HMI tags "Digitais"
   "Digitais_MB-01-YR" : Bool = PLC Digitais.MB-01-YR AT %DB300.DBX0.1, 1 s
   "Digitais_MB-01-YF" : Bool = PLC Digitais.MB-01-YF AT %DB300.DBX0.2, 1 s
   "Digitais_MB-01-YFF" : Bool = PLC Digitais.MB-01-YFF AT %DB300.DBX0.3, 1 s
   "Digitais_MB-01-MM" : Bool = PLC Digitais.MB-01-MM AT %DB300.DBX0.4, 1 s
   "Digitais_MB-01-MA" : Bool = PLC Digitais.MB-01-MA AT %DB300.DBX0.5, 1 s
   "Digitais_MB-01-EMER" : Bool = PLC Digitais.MB-01-EMER AT %DB300.DBX0.6, 1 s
   "Digitais_MB-01-MN" : Bool = PLC Digitais.MB-01-MN AT %DB300.DBX0.7, 1 s
   "Digitais_MB-01-ML" : Bool = PLC Digitais.MB-01-ML AT %DB300.DBX1.0, 1 s
   "Digitais_MB-01-YFI" : Bool = PLC Digitais.MB-01-YFI AT %DB300.DBX1.1, 1 s
   "Digitais_MB-01-YFA" : Bool = PLC Digitais.MB-01-YFA AT %DB300.DBX1.2, 1 s
   "Digitais_MB-01-YPTA" : Bool = PLC Digitais.MB-01-YPTA AT %DB300.DBX1.3, 1 s
   "Digitais_MB-01-HM" : Bool = PLC Digitais.MB-01-HM AT %DB300.DBX1.4, 1 s
   "Digitais_MB-01-RST" : Bool = PLC Digitais.MB-01-RST AT %DB300.DBX1.5, 1 s
   "Digitais_MB-01-INTRU" : Bool = PLC Digitais.MB-01-INTRU AT %DB300.DBX1.6, 1 s
   "Digitais_MB-01-YFB" : Bool = PLC Digitais.MB-01-YFB AT %DB300.DBX1.7, 1 s
   "Digitais_MB-02-YSH" : Bool = PLC Digitais.MB-02-YSH AT %DB300.DBX2.0, 1 s
   "Digitais_MB-02-YR" : Bool = PLC Digitais.MB-02-YR AT %DB300.DBX2.1, 1 s
   "Digitais_MB-02-YF" : Bool = PLC Digitais.MB-02-YF AT %DB300.DBX2.2, 1 s
   "Digitais_MB-02-YFF" : Bool = PLC Digitais.MB-02-YFF AT %DB300.DBX2.3, 1 s
   "Digitais_MB-02-MM" : Bool = PLC Digitais.MB-02-MM AT %DB300.DBX2.4, 1 s
   "Digitais_MB-02-MA" : Bool = PLC Digitais.MB-02-MA AT %DB300.DBX2.5, 1 s
   "Digitais_MB-02-EMER" : Bool = PLC Digitais.MB-02-EMER AT %DB300.DBX2.6, 1 s
   "Digitais_MB-02-MN" : Bool = PLC Digitais.MB-02-MN AT %DB300.DBX2.7, 1 s
   "Digitais_MB-02-ML" : Bool = PLC Digitais.MB-02-ML AT %DB300.DBX3.0, 1 s
   "Digitais_MB-02-YFI" : Bool = PLC Digitais.MB-02-YFI AT %DB300.DBX3.1, 1 s
   "Digitais_MB-02-YFA" : Bool = PLC Digitais.MB-02-YFA AT %DB300.DBX3.2, 1 s
   "Digitais_MB-02-YPTA" : Bool = PLC Digitais.MB-02-YPTA AT %DB300.DBX3.3, 1 s
   "Digitais_MB-02-HM" : Bool = PLC Digitais.MB-02-HM AT %DB300.DBX3.4, 1 s
   "Digitais_MB-02-RST" : Bool = PLC Digitais.MB-02-RST AT %DB300.DBX3.5, 1 s
   "Digitais_MB-02-INTRU" : Bool = PLC Digitais.MB-02-INTRU AT %DB300.DBX3.6, 1 s
   "Digitais_MB-02-YFB" : Bool = PLC Digitais.MB-02-YFB AT %DB300.DBX3.7, 1 s
   "Digitais_MB-03-YSH" : Bool = PLC Digitais.MB-03-YSH AT %DB300.DBX4.0, 1 s
   "Digitais_MB-03-YR" : Bool = PLC Digitais.MB-03-YR AT %DB300.DBX4.1, 1 s
   "Digitais_MB-03-YF" : Bool = PLC Digitais.MB-03-YF AT %DB300.DBX4.2, 1 s
   "Digitais_MB-03-YFF" : Bool = PLC Digitais.MB-03-YFF AT %DB300.DBX4.3, 1 s
   "Digitais_MB-03-MM" : Bool = PLC Digitais.MB-03-MM AT %DB300.DBX4.4, 1 s
   "Digitais_MB-03-MA" : Bool = PLC Digitais.MB-03-MA AT %DB300.DBX4.5, 1 s
   "Digitais_MB-03-EMER" : Bool = PLC Digitais.MB-03-EMER AT %DB300.DBX4.6, 1 s
   "Digitais_MB-03-MN" : Bool = PLC Digitais.MB-03-MN AT %DB300.DBX4.7, 1 s
   "Digitais_MB-03-ML" : Bool = PLC Digitais.MB-03-ML AT %DB300.DBX5.0, 1 s
   "Digitais_MB-03-YFI" : Bool = PLC Digitais.MB-03-YFI AT %DB300.DBX5.1, 1 s
   "Digitais_MB-03-YFA" : Bool = PLC Digitais.MB-03-YFA AT %DB300.DBX5.2, 1 s
   "Digitais_MB-03-YPTA" : Bool = PLC Digitais.MB-03-YPTA AT %DB300.DBX5.3, 1 s
   "Digitais_MB-03-HM" : Bool = PLC Digitais.MB-03-HM AT %DB300.DBX5.4, 1 s
   "Digitais_MB-03-RST" : Bool = PLC Digitais.MB-03-RST AT %DB300.DBX5.5, 1 s
   "Digitais_MB-03-INTRU" : Bool = PLC Digitais.MB-03-INTRU AT %DB300.DBX5.6, 1 s
   "Digitais_MB-03-YFB" : Bool = PLC Digitais.MB-03-YFB AT %DB300.DBX5.7, 1 s
   "Digitais_MB-04-YSH" : Bool = PLC Digitais.MB-04-YSH AT %DB300.DBX6.0, 1 s
   "Digitais_MB-04-YR" : Bool = PLC Digitais.MB-04-YR AT %DB300.DBX6.1, 1 s
   "Digitais_MB-04-YF" : Bool = PLC Digitais.MB-04-YF AT %DB300.DBX6.2, 1 s
   "Digitais_MB-04-YFF" : Bool = PLC Digitais.MB-04-YFF AT %DB300.DBX6.3, 1 s
   "Digitais_MB-04-MM" : Bool = PLC Digitais.MB-04-MM AT %DB300.DBX6.4, 1 s
   "Digitais_MB-04-MA" : Bool = PLC Digitais.MB-04-MA AT %DB300.DBX6.5, 1 s
   "Digitais_MB-04-EMER" : Bool = PLC Digitais.MB-04-EMER AT %DB300.DBX6.6, 1 s
   "Digitais_MB-04-MN" : Bool = PLC Digitais.MB-04-MN AT %DB300.DBX6.7, 1 s
   "Digitais_MB-04-ML" : Bool = PLC Digitais.MB-04-ML AT %DB300.DBX7.0, 1 s
   "Digitais_MB-04-YFI" : Bool = PLC Digitais.MB-04-YFI AT %DB300.DBX7.1, 1 s
   "Digitais_MB-04-YFA" : Bool = PLC Digitais.MB-04-YFA AT %DB300.DBX7.2, 1 s
   "Digitais_MB-04-YPTA" : Bool = PLC Digitais.MB-04-YPTA AT %DB300.DBX7.3, 1 s
   "Digitais_MB-04-HM" : Bool = PLC Digitais.MB-04-HM AT %DB300.DBX7.4, 1 s
   "Digitais_MB-04-RST" : Bool = PLC Digitais.MB-04-RST AT %DB300.DBX7.5, 1 s
   "Digitais_MB-04-INTRU" : Bool = PLC Digitais.MB-04-INTRU AT %DB300.DBX7.6, 1 s
   "Digitais_MB-04-YFB" : Bool = PLC Digitais.MB-04-YFB AT %DB300.DBX7.7, 1 s
   "Digitais_LIT_001-AL8" : Bool = PLC Digitais.LIT_001-AL8 AT %DB300.DBX8.0, 1 s
   "Digitais_LIT_001-AL9" : Bool = PLC Digitais.LIT_001-AL9 AT %DB300.DBX8.1, 1 s
   "Digitais_LIT_001-AL10" : Bool = PLC Digitais.LIT_001-AL10 AT %DB300.DBX8.2, 1 s
   "Digitais_LIT_001-AL11" : Bool = PLC Digitais.LIT_001-AL11 AT %DB300.DBX8.3, 1 s
   "Digitais_LIT_001-AL12" : Bool = PLC Digitais.LIT_001-AL12 AT %DB300.DBX8.4, 1 s
   "Digitais_LIT_001-AL13" : Bool = PLC Digitais.LIT_001-AL13 AT %DB300.DBX8.5, 1 s
   "Digitais_LIT_001-AL14" : Bool = PLC Digitais.LIT_001-AL14 AT %DB300.DBX8.6, 1 s
   "Digitais_LIT_001-AL15" : Bool = PLC Digitais.LIT_001-AL15 AT %DB300.DBX8.7, 1 s
   "Digitais_LIT_001-YHH" : Bool = PLC Digitais.LIT_001-YHH AT %DB300.DBX9.0, 1 s
   "Digitais_LIT_001-YH" : Bool = PLC Digitais.LIT_001-YH AT %DB300.DBX9.1, 1 s
   "Digitais_LIT_001-YL" : Bool = PLC Digitais.LIT_001-YL AT %DB300.DBX9.2, 1 s
   "Digitais_LIT_001-YLL" : Bool = PLC Digitais.LIT_001-YLL AT %DB300.DBX9.3, 1 s
   "Digitais_LIT_001-YFS" : Bool = PLC Digitais.LIT_001-YFS AT %DB300.DBX9.4, 1 s
   "Digitais_LIT_001-AL5" : Bool = PLC Digitais.LIT_001-AL5 AT %DB300.DBX9.5, 1 s
   "Digitais_LIT_001-AL6" : Bool = PLC Digitais.LIT_001-AL6 AT %DB300.DBX9.6, 1 s
   "Digitais_LIT_001-AL7" : Bool = PLC Digitais.LIT_001-AL7 AT %DB300.DBX9.7, 1 s
   "Digitais_PCM_EEE_EMER" : Bool = PLC Digitais.PCM_EEE_EMER AT %DB300.DBX10.0, 1 s
   "Digitais_PCM_EEE_K27" : Bool = PLC Digitais.PCM_EEE_K27 AT %DB300.DBX10.1, 1 s
   "Digitais_PCM_EEE_DISJ_LIG" : Bool = PLC Digitais.PCM_EEE_DISJ_LIG AT %DB300.DBX10.2, 1 s
   "Digitais_PCM_EEE_DISJ_DESLIG" : Bool = PLC Digitais.PCM_EEE_DISJ_DESLIG AT %DB300.DBX10.3, 1 s
   "Digitais_PCM_EEE_DISJ_YFAL" : Bool = PLC Digitais.PCM_EEE_DISJ_YFAL AT %DB300.DBX10.4, 1 s
   "Digitais_PCM_EEE_DISJ_FAL_GR" : Bool = PLC Digitais.PCM_EEE_DISJ_FAL_GR AT %DB300.DBX10.5, 1 s
   "Digitais_PCM_EEE_TR01_KA3" : Bool = PLC Digitais.PCM_EEE_TR01_KA3 AT %DB300.DBX10.6, 1 s
   "Digitais_PCM_EEE_TR01_KA4" : Bool = PLC Digitais.PCM_EEE_TR01_KA4 AT %DB300.DBX10.7, 1 s
   "Digitais_PCM_EEE_TR01_KA5" : Bool = PLC Digitais.PCM_EEE_TR01_KA5 AT %DB300.DBX11.0, 1 s
   "Digitais_PCM_EEE_INTRU" : Bool = PLC Digitais.PCM_EEE_INTRU AT %DB300.DBX11.1, 1 s
   "Digitais_PCM_EEE_RSERVA_0" : Bool = PLC Digitais.PCM_EEE_RSERVA_0 AT %DB300.DBX11.2, 1 s
   "Digitais_PCM_EEE_RSERVA_1" : Bool = PLC Digitais.PCM_EEE_RSERVA_1 AT %DB300.DBX11.3, 1 s
   "Digitais_PCM_EEE_RSERVA_2" : Bool = PLC Digitais.PCM_EEE_RSERVA_2 AT %DB300.DBX11.4, 1 s
   "Digitais_PCM_EEE_RSERVA_3" : Bool = PLC Digitais.PCM_EEE_RSERVA_3 AT %DB300.DBX11.5, 1 s
   "Digitais_PCM_EEE_RSERVA_4" : Bool = PLC Digitais.PCM_EEE_RSERVA_4 AT %DB300.DBX11.6, 1 s
   "Digitais_PCM_EEE_RSERVA_5" : Bool = PLC Digitais.PCM_EEE_RSERVA_5 AT %DB300.DBX11.7, 1 s
   "Digitais_QGBT_EMER" : Bool = PLC Digitais.QGBT_EMER AT %DB300.DBX12.0, 1 s
   "Digitais_QGBT_K27" : Bool = PLC Digitais.QGBT_K27 AT %DB300.DBX12.1, 1 s
   "Digitais_QGBT_DJL" : Bool = PLC Digitais.QGBT_DJL AT %DB300.DBX12.2, 1 s
   "Digitais_QGBT_DJD" : Bool = PLC Digitais.QGBT_DJD AT %DB300.DBX12.3, 1 s
   "Digitais_QGBT_DJYFAL" : Bool = PLC Digitais.QGBT_DJYFAL AT %DB300.DBX12.4, 1 s
   "Digitais_QGBT_INTRU" : Bool = PLC Digitais.QGBT_INTRU AT %DB300.DBX12.5, 1 s
   "Digitais_QGBT_RESERVA_0" : Bool = PLC Digitais.QGBT_RESERVA_0 AT %DB300.DBX12.6, 1 s
   "Digitais_QGBT_RESERVA_1" : Bool = PLC Digitais.QGBT_RESERVA_1 AT %DB300.DBX12.7, 1 s
   "Digitais_QGBT_RESERVA_2" : Bool = PLC Digitais.QGBT_RESERVA_2 AT %DB300.DBX13.0, 1 s
   "Digitais_QGBT_RESERVA_3" : Bool = PLC Digitais.QGBT_RESERVA_3 AT %DB300.DBX13.1, 1 s
   "Digitais_QGBT_RESERVA_4" : Bool = PLC Digitais.QGBT_RESERVA_4 AT %DB300.DBX13.2, 1 s
   "Digitais_QGBT_RESERVA_5" : Bool = PLC Digitais.QGBT_RESERVA_5 AT %DB300.DBX13.3, 1 s
   "Digitais_QGBT_RESERVA_6" : Bool = PLC Digitais.QGBT_RESERVA_6 AT %DB300.DBX13.4, 1 s
   "Digitais_QGBT_RESERVA_7" : Bool = PLC Digitais.QGBT_RESERVA_7 AT %DB300.DBX13.5, 1 s
   "Digitais_QGBT_RESERVA_8" : Bool = PLC Digitais.QGBT_RESERVA_8 AT %DB300.DBX13.6, 1 s
   "Digitais_QGBT_RESERVA_9" : Bool = PLC Digitais.QGBT_RESERVA_9 AT %DB300.DBX13.7, 1 s
   "Digitais_LSL_001" : Bool = PLC Digitais.LSL_001 AT %DB300.DBX14.0, 1 s
   "Digitais_LSH_001" : Bool = PLC Digitais.LSH_001 AT %DB300.DBX14.1, 1 s
   "Digitais_LSL_002" : Bool = PLC Digitais.LSL_002 AT %DB300.DBX14.2, 1 s
   "Digitais_LSH_002" : Bool = PLC Digitais.LSH_002 AT %DB300.DBX14.3, 1 s
   "Digitais_LS_RESERVA_0" : Bool = PLC Digitais.LS_RESERVA_0 AT %DB300.DBX14.4, 1 s
   "Digitais_LS_RESERVA_1" : Bool = PLC Digitais.LS_RESERVA_1 AT %DB300.DBX14.5, 1 s
   "Digitais_LS_RESERVA_2" : Bool = PLC Digitais.LS_RESERVA_2 AT %DB300.DBX14.6, 1 s
   "Digitais_LS_RESERVA_3" : Bool = PLC Digitais.LS_RESERVA_3 AT %DB300.DBX14.7, 1 s
   "Digitais_LS_RESERVA_4" : Bool = PLC Digitais.LS_RESERVA_4 AT %DB300.DBX15.0, 1 s
   "Digitais_LS_RESERVA_5" : Bool = PLC Digitais.LS_RESERVA_5 AT %DB300.DBX15.1, 1 s
   "Digitais_LS_RESERVA_6" : Bool = PLC Digitais.LS_RESERVA_6 AT %DB300.DBX15.2, 1 s
   "Digitais_LS_RESERVA_7" : Bool = PLC Digitais.LS_RESERVA_7 AT %DB300.DBX15.3, 1 s
   "Digitais_LS_RESERVA_8" : Bool = PLC Digitais.LS_RESERVA_8 AT %DB300.DBX15.4, 1 s
   "Digitais_LS_RESERVA_9" : Bool = PLC Digitais.LS_RESERVA_9 AT %DB300.DBX15.5, 1 s
   "Digitais_LS_RESERVA_10" : Bool = PLC Digitais.LS_RESERVA_10 AT %DB300.DBX15.6, 1 s
   "Digitais_LS_RESERVA_11" : Bool = PLC Digitais.LS_RESERVA_11 AT %DB300.DBX15.7, 1 s
   "Digitais_PCE_EEE_INTRU" : Bool = PLC Digitais.PCE_EEE_INTRU AT %DB300.DBX16.0, 1 s
   "Digitais_PCE_EEE_UPS_ALM" : Bool = PLC Digitais.PCE_EEE_UPS_ALM AT %DB300.DBX16.1, 1 s
   "Digitais_PCE_EEE_UPS_FE" : Bool = PLC Digitais.PCE_EEE_UPS_FE AT %DB300.DBX16.2, 1 s
   "Digitais_PCE_EEE_UPS_CHAR" : Bool = PLC Digitais.PCE_EEE_UPS_CHAR AT %DB300.DBX16.3, 1 s
   "Digitais_PCM-E-CF-01-P100-YFC" : Bool = PLC Digitais.PCM-E-CF-01-P100-YFC AT %DB300.DBX16.4, 1 s
   "Digitais_QGBT-AUX-01-P100-YFC" : Bool = PLC Digitais.QGBT-AUX-01-P100-YFC AT %DB300.DBX16.5, 1 s

HMI tags "Setpoints"
   "SETPOINTS_MB-01-SP" : Real = PLC SETPOINTS.MB-01-SP AT %DB305.DBD0, 1 s
   "SETPOINTS_MB-02-SP" : Real = PLC SETPOINTS.MB-02-SP AT %DB305.DBD4, 1 s
   "SETPOINTS_MB-03-SP" : Real = PLC SETPOINTS.MB-03-SP AT %DB305.DBD8, 1 s
   "SETPOINTS_MB-04-SP" : Real = PLC SETPOINTS.MB-04-SP AT %DB305.DBD12, 1 s
   "SETPOINTS_LIT_001-SPHH" : Real = PLC SETPOINTS.LIT_001-SPHH AT %DB305.DBD16, 1 s
   "SETPOINTS_LIT_001-SPH" : Real = PLC SETPOINTS.LIT_001-SPH AT %DB305.DBD20, 1 s
   "SETPOINTS_LIT_001-SPL" : Real = PLC SETPOINTS.LIT_001-SPL AT %DB305.DBD24, 1 s
   "SETPOINTS_LIT_001-SPLL" : Real = PLC SETPOINTS.LIT_001-SPLL AT %DB305.DBD28, 1 s
   "SETPOINTS_LIT_001-SPM" : Real = PLC SETPOINTS.LIT_001-SPM AT %DB305.DBD32, 1 s
   "SETPOINTS_LIT_001-SPC" : Real = PLC SETPOINTS.LIT_001-SPC AT %DB305.DBD36, 1 s
   "SETPOINTS_LIT-001-P" : Real = PLC SETPOINTS.LIT-001-P AT %DB305.DBD40, 1 s
   "SETPOINTS_SP_NVL_MIN" : Real = PLC SETPOINTS.SP_NVL_MIN AT %DB305.DBD44, 1 s
   "SETPOINTS_MB-P-SP-DL" : Real = PLC SETPOINTS.MB-P-SP-DL AT %DB305.DBD48, 1 s
   "SETPOINTS_MB-P-SP-L" : Real = PLC SETPOINTS.MB-P-SP-L AT %DB305.DBD52, 1 s
   "SETPOINTS_MB-C1-SP-DL" : Real = PLC SETPOINTS.MB-C1-SP-DL AT %DB305.DBD56, 1 s
   "SETPOINTS_MB-C1-SP-L" : Real = PLC SETPOINTS.MB-C1-SP-L AT %DB305.DBD60, 1 s
   "SETPOINTS_MB-C2-SP-DL" : Real = PLC SETPOINTS.MB-C2-SP-DL AT %DB305.DBD64, 1 s
   "SETPOINTS_MB-C2-SP-L" : Real = PLC SETPOINTS.MB-C2-SP-L AT %DB305.DBD68, 1 s
   "SETPOINTS_MB-C3-SP-DL" : Real = PLC SETPOINTS.MB-C3-SP-DL AT %DB305.DBD72, 1 s
   "SETPOINTS_MB-C3-SP-L" : Real = PLC SETPOINTS.MB-C3-SP-L AT %DB305.DBD76, 1 s

HMI tags "Variaveis"
   "VARIAVEIS_MB-01-YST" : Real = PLC VARIAVEIS.MB-01-YST AT %DB304.DBD0, 1 s
   "VARIAVEIS_MB-01-YIT" : Real = PLC VARIAVEIS.MB-01-YIT AT %DB304.DBD4, 1 s
   "VARIAVEIS_MB-02-YIT" : Real = PLC VARIAVEIS.MB-02-YIT AT %DB304.DBD8, 1 s
   "VARIAVEIS_MB-02-YST" : Real = PLC VARIAVEIS.MB-02-YST AT %DB304.DBD12, 1 s
   "VARIAVEIS_MB-03-YIT" : Real = PLC VARIAVEIS.MB-03-YIT AT %DB304.DBD16, 1 s
   "VARIAVEIS_MB-03-YST" : Real = PLC VARIAVEIS.MB-03-YST AT %DB304.DBD20, 1 s
   "VARIAVEIS_MB-04-YIT" : Real = PLC VARIAVEIS.MB-04-YIT AT %DB304.DBD24, 1 s
   "VARIAVEIS_MB-04-YST" : Real = PLC VARIAVEIS.MB-04-YST AT %DB304.DBD28, 1 s
   "VARIAVEIS_LIT_001" : Real = PLC VARIAVEIS.LIT_001 AT %DB304.DBD32, 1 s
   "VARIAVEIS_LIT_001-P" : Real = PLC VARIAVEIS.LIT_001-P AT %DB304.DBD36, 1 s
   "VARIAVEIS_PCM-E-CF-01-04-P100-ETRS" : Real = PLC VARIAVEIS.PCM-E-CF-01-04-P100-ETRS AT %DB304.DBD40, 1 s
   "VARIAVEIS_PCM-E-CF-01-04-P100-ETST" : Real = PLC VARIAVEIS.PCM-E-CF-01-04-P100-ETST AT %DB304.DBD44, 1 s
   "VARIAVEIS_PCM-E-CF-01-04-P100-ETTR" : Real = PLC VARIAVEIS.PCM-E-CF-01-04-P100-ETTR AT %DB304.DBD48, 1 s
   "VARIAVEIS_PCM-E-CF-01-04-P100-ITR" : Real = PLC VARIAVEIS.PCM-E-CF-01-04-P100-ITR AT %DB304.DBD52, 1 s
   "VARIAVEIS_PCM-E-CF-01-04-P100-ITS" : Real = PLC VARIAVEIS.PCM-E-CF-01-04-P100-ITS AT %DB304.DBD56, 1 s
   "VARIAVEIS_PCM-E-CF-01-04-P100-ITT" : Real = PLC VARIAVEIS.PCM-E-CF-01-04-P100-ITT AT %DB304.DBD60, 1 s
   "VARIAVEIS_PCM-E-CF-01-04-P100-JPT" : Real = PLC VARIAVEIS.PCM-E-CF-01-04-P100-JPT AT %DB304.DBD64, 1 s
   "VARIAVEIS_PCM-E-CF-01-04-P100-JQT" : Real = PLC VARIAVEIS.PCM-E-CF-01-04-P100-JQT AT %DB304.DBD68, 1 s
   "VARIAVEIS_PCM-E-CF-01-04-P100-JST" : Real = PLC VARIAVEIS.PCM-E-CF-01-04-P100-JST AT %DB304.DBD72, 1 s
   "VARIAVEIS_PCM-E-CF-01-04-P100-FP" : Real = PLC VARIAVEIS.PCM-E-CF-01-04-P100-FP AT %DB304.DBD76, 1 s
   "VARIAVEIS_QGBT-AUX-01-P100-ETRS" : Real = PLC VARIAVEIS.QGBT-AUX-01-P100-ETRS AT %DB304.DBD80, 1 s
   "VARIAVEIS_QGBT-AUX-01-P100-ETST" : Real = PLC VARIAVEIS.QGBT-AUX-01-P100-ETST AT %DB304.DBD84, 1 s
   "VARIAVEIS_QGBT-AUX-01-P100-ETTR" : Real = PLC VARIAVEIS.QGBT-AUX-01-P100-ETTR AT %DB304.DBD88, 1 s
   "VARIAVEIS_QGBT-AUX-01-P100-ITR" : Real = PLC VARIAVEIS.QGBT-AUX-01-P100-ITR AT %DB304.DBD92, 1 s
   "VARIAVEIS_QGBT-AUX-01-P100-ITS" : Real = PLC VARIAVEIS.QGBT-AUX-01-P100-ITS AT %DB304.DBD96, 1 s
   "VARIAVEIS_QGBT-AUX-01-P100-ITT" : Real = PLC VARIAVEIS.QGBT-AUX-01-P100-ITT AT %DB304.DBD100, 1 s
   "VARIAVEIS_QGBT-AUX-01-P100-JPT" : Real = PLC VARIAVEIS.QGBT-AUX-01-P100-JPT AT %DB304.DBD104, 1 s
   "VARIAVEIS_QGBT-AUX-01-P100-JQT" : Real = PLC VARIAVEIS.QGBT-AUX-01-P100-JQT AT %DB304.DBD108, 1 s
   "VARIAVEIS_QGBT-AUX-01-P100-JST" : Real = PLC VARIAVEIS.QGBT-AUX-01-P100-JST AT %DB304.DBD112, 1 s
   "VARIAVEIS_QGBT-AUX-01-P100-FP" : Real = PLC VARIAVEIS.QGBT-AUX-01-P100-FP AT %DB304.DBD116, 1 s

HMI tags "STATUS"
   "STATUS_MB-01-YSP" : Bool = PLC STATUS.MB-01-YSP AT %DB302.DBX0.6, 1 s
   "STATUS_MB-02-YSP" : Bool = PLC STATUS.MB-02-YSP AT %DB302.DBX0.7, 1 s
   "STATUS_MB-03-YSP" : Bool = PLC STATUS.MB-03-YSP AT %DB302.DBX1.1, 1 s
   "STATUS_MB-01-YC1" : Bool = PLC STATUS.MB-01-YC1 AT %DB302.DBX1.2, 1 s
   "STATUS_MB-02-YC1" : Bool = PLC STATUS.MB-02-YC1 AT %DB302.DBX1.3, 1 s
   "STATUS_MB-03-YC1" : Bool = PLC STATUS.MB-03-YC1 AT %DB302.DBX1.5, 1 s
   "STATUS_MB-01-YC2" : Bool = PLC STATUS.MB-01-YC2 AT %DB302.DBX1.6, 1 s
   "STATUS_MB-02-YC2" : Bool = PLC STATUS.MB-02-YC2 AT %DB302.DBX1.7, 1 s
   "STATUS_MB-03-YC2" : Bool = PLC STATUS.MB-03-YC2 AT %DB302.DBX2.1, 1 s
   "STATUS_MB-04-YSP" : Bool = PLC STATUS.MB-04-YSP AT %DB302.DBX1.0, 1 s
   "STATUS_MB-04-YC1" : Bool = PLC STATUS.MB-04-YC1 AT %DB302.DBX1.4, 1 s
   "STATUS_MB-04-YC2" : Bool = PLC STATUS.MB-04-YC2 AT %DB302.DBX2.0, 1 s

discrete alarms
   1: 'Elevatoria principal 1 falha', class Errors, trigger "ALM0" bit 10
   2: 'Elevatoria principal 1 falta de fase', class Errors, trigger "ALM0" bit 11
   3: 'Elevatoria principal 1 emergencia', class Errors, trigger "ALM0" bit 14
   5: 'Elevatoria principal 1 com falha no inversor', class Errors, trigger "ALM0" bit 1
   6: 'Elevatoria principal 1 com falha no acionamento', class Errors, trigger "ALM0" bit 2
   7: 'Elevatoria principal 1 com proteção térmica atuada', class Errors, trigger "ALM0" bit 3
   8: 'Elevatoria principal 1 intrusão no painel', class Errors, trigger "ALM0" bit 6
   9: 'Elevatoria principal 1 defeito na bomba', class Errors, trigger "ALM0" bit 7
   10: 'Elevatoria principal 2 falha', class Errors, trigger "ALM2" bit 10
   11: 'Elevatoria principal 2 falta de fase', class Errors, trigger "ALM2" bit 11
   12: 'Elevatoria principal 2 emergencia', class Errors, trigger "ALM2" bit 14
   14: 'Elevatoria principal 2 com falha no inversor', class Errors, trigger "ALM2" bit 1
   15: 'Elevatoria principal 2 com falha no acionamento', class Errors, trigger "ALM2" bit 2
   16: 'Elevatoria principal 2 com proteção térmica atuada', class Errors, trigger "ALM2" bit 3
   17: 'Elevatoria principal 2 intrusão no painel', class Errors, trigger "ALM2" bit 6
   18: 'Elevatoria principal 2 defeito na bomba', class Errors, trigger "ALM2" bit 7
   19: 'Elevatoria principal 3 falha', class Errors, trigger "ALM4" bit 10
   20: 'Elevatoria principal 3 falta de fase', class Errors, trigger "ALM4" bit 11
   21: 'Elevatoria principal 3 emergencia', class Errors, trigger "ALM4" bit 14
   23: 'Elevatoria principal 3 com falha no inversor', class Errors, trigger "ALM4" bit 1
   24: 'Elevatoria principal 3 com falha no acionamento', class Errors, trigger "ALM4" bit 2
   25: 'Elevatoria principal 3 com proteção térmica atuada', class Errors, trigger "ALM4" bit 3
   26: 'Elevatoria principal 3 intrusão no painel', class Errors, trigger "ALM4" bit 6
   27: 'Elevatoria principal 3 defeito na bomba', class Errors, trigger "ALM4" bit 7
   28: 'Elevatoria principal 4 falha', class Errors, trigger "ALM6" bit 10
   29: 'Elevatoria principal 4 falta de fase', class Errors, trigger "ALM6" bit 11
   30: 'Elevatoria principal 4 emergencia', class Errors, trigger "ALM6" bit 14
   32: 'Elevatoria principal 4 com falha no inversor', class Errors, trigger "ALM6" bit 1
   33: 'Elevatoria principal 4 com falha no acionamento', class Errors, trigger "ALM6" bit 2
   34: 'Elevatoria principal 4 com proteção térmica atuada', class Errors, trigger "ALM6" bit 3
   35: 'Elevatoria principal 4 intrusão no painel', class Errors, trigger "ALM6" bit 6
   36: 'Elevatoria principal 4 defeito na bomba', class Errors, trigger "ALM6" bit 7
   37: 'Alarme de nível muito alto do tanque', class Errors, trigger "ALM8" bit 0
   38: 'Alarme de nível alto do tanque', class Errors, trigger "ALM8" bit 1
   39: 'Alarme de nível baixo do tanque', class Errors, trigger "ALM8" bit 2
   40: 'Alarme de nível muito baixo do tanque', class Errors, trigger "ALM8" bit 3
   41: 'Transmissor de nível do tanque com falha de sinal', class Errors, trigger "ALM8" bit 4
   42: 'PCM-E-CF-01-04 BOTAO DE EMERGENCIA - ATUADO', class Errors, trigger "ALM10" bit 8
   43: 'PCM-E-CF-01-04 RELE DE PROTECAO FUNCAO 27 - ATUADO', class Errors, trigger "ALM10" bit 9
   44: 'PCM-E-CF-01-04 DISJUNTOR GERAL STATUS - FALHA', class Errors, trigger "ALM10" bit 12
   45: 'PCM-E-CF-01-04 FALHA GERAL ATUADO', class Errors, trigger "ALM10" bit 13
   46: 'PCM-E-CF-01-04 TRANSFORMADOR -TR-01 ALARME TEMP 150°', class Errors, trigger "ALM10" bit 14
   47: 'PCM-E-CF-01-04 TRANSFORMADOR -TR-01 ALARME TEMP 155°', class Errors, trigger "ALM10" bit 15
   48: 'PCM-E-CF-01-04 TRANSFORMADOR -TR-01 FALHA PROTECAO', class Errors, trigger "ALM10" bit 0
   49: 'PCM-E-CF-01-04 INTRUSAO NO PAINEL (COLUNA 01~04)', class Errors, trigger "ALM10" bit 1
   50: 'QGBT-AUX-01 BOTAO DE EMERGENCIA ATUADO', class Errors, trigger "ALM12" bit 8
   51: 'QGBT-AUX-01 RELE DE PROTECAO FUNCAO 27/59 ATUADO', class Errors, trigger "ALM12" bit 9
   52: 'QGBT-AUX-01 DISJUNTOR GERAL FALHA - TRIP', class Errors, trigger "ALM12" bit 12
   53: 'QGBT-AUX-01 INTRUSAO NO PAINEL', class Errors, trigger "ALM12" bit 13
   54: 'INTRUSAO NO PAINEL', class Errors, trigger "ALM16" bit 8
   55: 'UPS EM ALARME FALHA NA BATERIA', class Errors, trigger "ALM16" bit 9
   56: 'UPS EM OPERACAO FALTA DE ENERGIA', class Errors, trigger "ALM16" bit 10
   57: 'UPS EM ALARME BATERIA CARREGADA', class Errors, trigger "ALM16" bit 11

screen "EEEB" 800x480, template "Template_1"
   GraphicView "Template_Graphic view_3" at 143,92 size 589x312; Picture "EEEB_2"
   Bar "Bar_1" at 679,137 size 57x267; MinimumValue 0; MaximumValue 100
      ProcessValue <- "VARIAVEIS_LIT_001-P"
   GraphicView "Graphic view_1" at 280,337 size 47x47; Picture "Submersa_vm"
      Visibility <- "Digitais_MB-01-YSH"
   GraphicView "Graphic view_2" at 280,337 size 47x47; Picture "Submersa_am"
      Visibility <- "Digitais_MB-01-YF"
   GraphicView "Graphic view_3" at 280,337 size 47x47; Picture "Submersa_azul"
      Visibility <- "COMANDOS_MB-01-HS7"
   GraphicView "Graphic view_4" at 395,337 size 47x47; Picture "Submersa_vm"
      Visibility <- "Digitais_MB-02-YSH"
   GraphicView "Graphic view_5" at 395,337 size 47x47; Picture "Submersa_am"
      Visibility <- "Digitais_MB-02-YF"
   GraphicView "Graphic view_6" at 395,337 size 47x47; Picture "Submersa_azul"
      Visibility <- "COMANDOS_MB-02-HS7"
   GraphicView "Graphic view_7" at 510,337 size 47x47; Picture "Submersa_vm"
      Visibility <- "Digitais_MB-03-YSH"
   GraphicView "Graphic view_8" at 510,337 size 47x47; Picture "Submersa_am"
      Visibility <- "Digitais_MB-03-YF"
   GraphicView "Graphic view_9" at 510,337 size 47x47; Picture "Submersa_azul"
      Visibility <- "COMANDOS_MB-03-HS7"
   TextField "Text field_1" at 286,384 size 29x14; Text 'MB-01'
   TextField "Text field_2" at 403,384 size 29x14; Text 'MB-02'
   TextField "Text field_3" at 517,384 size 29x14; Text 'MB-03'
   TextField "Text field_4" at 248,328 size 25x16; Text 'AUT'
      Visibility <- "COMANDOS_MB-01-HS1"
   TextField "Text field_5" at 248,345 size 25x16; Text 'REM'
      Visibility <- "Digitais_MB-01-YR"
   TextField "Text field_6" at 296,322 size 25x16; Text 'P'
      Visibility <- "STATUS_MB-01-YSP"
   TextField "Text field_7" at 296,322 size 25x16; Text 'C1'
      Visibility <- "STATUS_MB-01-YC1"
   TextField "Text field_8" at 296,322 size 25x16; Text 'C2'
      Visibility <- "STATUS_MB-01-YC2"
   IOField "I/O field_3" at 222,363 size 54x17; FormatPattern 99.9; Unit  HZ
      ProcessValue <- "VARIAVEIS_MB-01-YST"
   IOField "I/O field_4" at 223,380 size 55x17; FormatPattern 999.9; Unit  A
      ProcessValue <- "VARIAVEIS_MB-01-YIT"
   TextField "Text field_9" at 364,328 size 25x16; Text 'AUT'
      Visibility <- "COMANDOS_MB-02-HS1"
   TextField "Text field_10" at 364,345 size 25x16; Text 'REM'
      Visibility <- "Digitais_MB-02-YR"
   TextField "Text field_11" at 412,322 size 25x16; Text 'P'
      Visibility <- "STATUS_MB-02-YSP"
   TextField "Text field_12" at 412,322 size 25x16; Text 'C1'
      Visibility <- "STATUS_MB-02-YC1"
   TextField "Text field_13" at 412,322 size 25x16; Text 'C2'
      Visibility <- "STATUS_MB-02-YC2"
   IOField "I/O field_5" at 338,363 size 54x17; FormatPattern 99.9; Unit  HZ
      ProcessValue <- "VARIAVEIS_MB-02-YST"
   IOField "I/O field_6" at 339,380 size 55x17; FormatPattern 999.9; Unit  A
      ProcessValue <- "VARIAVEIS_MB-02-YIT"
   TextField "Text field_14" at 478,328 size 25x16; Text 'AUT'
      Visibility <- "COMANDOS_MB-03-HS1"
   TextField "Text field_15" at 478,345 size 25x16; Text 'REM'
      Visibility <- "Digitais_MB-03-YR"
   TextField "Text field_16" at 526,322 size 25x16; Text 'P'
      Visibility <- "STATUS_MB-03-YSP"
   TextField "Text field_17" at 526,322 size 25x16; Text 'C1'
      Visibility <- "STATUS_MB-03-YC1"
   TextField "Text field_18" at 526,322 size 25x16; Text 'C2'
      Visibility <- "STATUS_MB-03-YC2"
   IOField "I/O field_7" at 452,363 size 54x17; FormatPattern 99.9; Unit  HZ
      ProcessValue <- "VARIAVEIS_MB-03-YST"
   IOField "I/O field_8" at 453,380 size 55x17; FormatPattern 999.9; Unit  A
      ProcessValue <- "VARIAVEIS_MB-03-YIT"
   IOField "I/O field_14" at 738,164 size 59x17; FormatPattern 99.99; Unit  m
      ProcessValue <- "VARIAVEIS_LIT_001"
      Appearance <- "Digitais_LIT_001-YFS"
   IOField "I/O field_17" at 738,180 size 59x17; FormatPattern 999.9; Unit  %
      ProcessValue <- "VARIAVEIS_LIT_001-P"
      Appearance <- "Digitais_LIT_001-YFS"
   TextField "Text field_19" at 772,148 size 25x16; Text 'HH'
      Visibility <- "Digitais_LIT_001-YHH"
   TextField "Text field_20" at 738,148 size 25x16; Text 'LL'
      Visibility <- "Digitais_LIT_001-YLL"
   TextField "Text field_21" at 738,197 size 25x16; Text 'L'
      Visibility <- "Digitais_LIT_001-YL"
   TextField "Text field_22" at 772,197 size 25x16; Text 'H'
      Visibility <- "Digitais_LIT_001-YH"
   Button "Button_5" at 332,10 size 96x32; TextOff 'pause loop'
      on Click: InvertBit("pause")
      Appearance <- "pause"
   IOField "I/O field_18" at 352,48 size 59x17; FormatPattern s99999
      ProcessValue <- "DIVERSOS_Looping"
      Visibility <- "pause"
   IOField "I/O field_1" at 567,363 size 54x17; FormatPattern 99.9; Unit  HZ
      ProcessValue <- "VARIAVEIS_MB-04-YST"
   IOField "I/O field_2" at 568,380 size 55x17; FormatPattern 999.9; Unit  A
      ProcessValue <- "VARIAVEIS_MB-04-YIT"
   TextField "Text field_23" at 646,322 size 25x16; Text 'P'
      Visibility <- "STATUS_MB-04-YSP"
   TextField "Text field_24" at 646,322 size 25x16; Text 'C1'
      Visibility <- "STATUS_MB-04-YC1"
   TextField "Text field_25" at 646,322 size 25x16; Text 'C2'
      Visibility <- "STATUS_MB-04-YC2"
   TextField "Text field_26" at 596,328 size 25x16; Text 'AUT'
      Visibility <- "COMANDOS_MB-04-HS1"
   TextField "Text field_27" at 596,345 size 25x16; Text 'REM'
      Visibility <- "Digitais_MB-04-YR"
   TextField "Text field_28" at 631,384 size 29x14; Text 'MB-04'
   GraphicView "Graphic view_10" at 624,337 size 47x47; Picture "Submersa_vm"
      Visibility <- "Digitais_MB-04-YSH"
   GraphicView "Graphic view_11" at 624,337 size 47x47; Picture "Submersa_am"
      Visibility <- "Digitais_MB-04-YF"
   GraphicView "Graphic view_12" at 624,337 size 47x47; Picture "Submersa_azul"
      Visibility <- "COMANDOS_MB-04-HS7"
   TextField "Text field_29" at 175,148 size 25x16; Text 'HH'
      Visibility <- "Digitais_LSH_002"
   TextField "Text field_30" at 175,378 size 25x16; Text 'LL'
      Visibility <- "Digitais_LSL_002"
   TextField "Text field_31" at 175,337 size 25x16; Text 'L'
      Visibility <- "Digitais_LSL_001"
   TextField "Text field_32" at 175,189 size 25x16; Text 'H'
      Visibility <- "Digitais_LSH_001"
   TextField "Text field_33" at 216,310 size 65x18; Text 'Manuteção'
      Visibility <- "Digitais_MB-01-MM"
   TextField "Text field_34" at 249,310 size 32x18; Text 'Local'
      Visibility <- "Digitais_MB-01-ML"
   TextField "Text field_35" at 217,310 size 64x18; Text 'Emegência'
      Visibility <- "Digitais_MB-01-EMER"
   TextField "Text field_36" at 331,310 size 65x18; Text 'Manuteção'
      Visibility <- "Digitais_MB-02-MM"
   TextField "Text field_37" at 364,310 size 32x18; Text 'Local'
      Visibility <- "Digitais_MB-02-ML"
   TextField "Text field_38" at 332,310 size 64x18; Text 'Emegência'
      Visibility <- "Digitais_MB-02-EMER"
   TextField "Text field_39" at 446,310 size 65x18; Text 'Manuteção'
      Visibility <- "Digitais_MB-03-MM"
   TextField "Text field_40" at 479,310 size 32x18; Text 'Local'
      Visibility <- "Digitais_MB-03-ML"
   TextField "Text field_41" at 447,310 size 64x18; Text 'Emegência'
      Visibility <- "Digitais_MB-03-EMER"
   TextField "Text field_42" at 561,310 size 65x18; Text 'Manuteção'
      Visibility <- "Digitais_MB-04-MM"
   TextField "Text field_43" at 594,310 size 32x18; Text 'Local'
      Visibility <- "Digitais_MB-04-ML"
   TextField "Text field_44" at 562,310 size 64x18; Text 'Emegência'
      Visibility <- "Digitais_MB-04-EMER"
   TextField "Text field_45" at 391,406 size 138x22; Text 'Emegência Acionado'
      Visibility <- "Digitais_PCM_EEE_EMER"

Template "Template_1" 800x480
   Button "Exit" at 724,444 size 50x36; TextOn 'Exit'; TextOff 'Exit'; PictureOn "ExitRuntime_KTP400_Basic_PN_TR"; PictureOff "SB_ExitRuntime_80x60_256c"
      on Release: StopRuntime(0)
   Button "Alarms" at 524,444 size 50x36; TextOn 'Alarms'; TextOff 'Alarms'; PictureOn "AlarmDisplay_KTP400_Basic_PN_TR"; PictureOff "AlarmDisplay_KTP400_Basic_PN_TR"
      on Release: function_ef3f5d25("Alarm window_1", -1)
   SymbolicIOField "Symbolic_IO_Field_Screen" at 185,7 size 510x49; TextOn '1'; TextOff '0'; TextList "TextList_ScreenNames"
      on Change: ActivateScreenByNumber("Tag_ScreenNumber", 0)
      ProcessValue <- "Tag_ScreenNumber"
   DateTimeField "HmiScreenItemData" at 695,29 size 102x22
   DateTimeField "HmiScreenItemData_1" at 686,5 size 111x22
   Group "Group" at 0,0 size 179x67; Picture "consbem"
   Button "Start screen_1" at 26,444 size 50x36; TextOn 'EEEB / Start screen'; TextOff 'EEEB / Start screen'; PictureOn "NavigateHome_KTP400_Basic_PN_TR"; PictureOff "NavigateHome_KTP400_Basic_PN_TR"
      on Release: ActivateScreen("EEEB", 1)
   Button "Start screen_2" at 125,444 size 50x36; TextOn 'Ajustes / Start screen'; TextOff 'Ajustes / Start screen'; PictureOn "NavigateHome_KTP400_Basic_PN_TR"; PictureOff "NavigateHome_KTP400_Basic_PN_TR"
      on Release: ActivateScreen("Ajustes", 1)
   Button "Start screen_3" at 226,444 size 50x36; TextOn 'Comando / Start screen'; TextOff 'Comando / Start screen'; PictureOn "NavigateHome_KTP400_Basic_PN_TR"; PictureOff "NavigateHome_KTP400_Basic_PN_TR"
      on Release: ActivateScreen("Comandos", 1)
   Button "Start screen_4" at 328,444 size 50x36; TextOn 'PID / Start screen'; TextOff 'PID / Start screen'; PictureOn "NavigateHome_KTP400_Basic_PN_TR"; PictureOff "NavigateHome_KTP400_Basic_PN_TR"
      on Release: ActivateScreen("PID", 1)
   Button "Start screen_5" at 426,444 size 50x36; TextOn 'Monitor. / Start screen'; TextOff 'Monitor. / Start screen'; PictureOn "NavigateHome_KTP400_Basic_PN_TR"; PictureOff "NavigateHome_KTP400_Basic_PN_TR"
      on Release: ActivateScreen("Monitoramento", 1)
   Softkey "Softkey_F1" at 0,0 size 0x0
      on KeyUp: ActivateScreen("EEEB", 0)
   Softkey "Softkey_F2" at 0,0 size 0x0
      on KeyUp: ActivateScreen("Ajustes", 1)
   Softkey "Softkey_F3" at 0,0 size 0x0
      on KeyUp: ActivateScreen("Comandos", 0)
   Softkey "Softkey_F4" at 0,0 size 0x0
      on KeyUp: ActivateScreen("PID", 1)
   GraphicView "Template_Graphic view_2" at 60,0 size 60x67; Picture "Consbem_novo"
   GraphicView "Template_Graphic view_3" at 119,0 size 60x67; Picture "logo-saae-header"
   GraphicView "Template_Graphic view_4" at 0,0 size 60x67; Picture "logo cápua"
   Softkey "Softkey_F5" at 0,0 size 0x0
      on KeyUp: ActivateScreen("Monitoramento", 0)
   Softkey "Softkey_F6" at 0,0 size 0x0
      on KeyUp: function_ef3f5d25("Alarm window_1", -1)

screen "Monitoramento" 800x480, template "Template_1"
   IOField "I/O field_9" at 649,330 size 71x17; FormatPattern 999.99; Unit  kW
      ProcessValue <- "VARIAVEIS_QGBT-AUX-01-P100-JPT"
      Appearance <- "Digitais_LIT_001-YFS"
   TextField "Text field_14" at 607,295 size 78x23; Text 'Potências'
   TextField "Text field_15" at 604,327 size 40x20; Text 'Ativa'
   IOField "I/O field_10" at 649,352 size 71x17; FormatPattern 999.99; Unit  KVA
      ProcessValue <- "VARIAVEIS_QGBT-AUX-01-P100-JST"
      Appearance <- "Digitais_LIT_001-YFS"
   TextField "Text field_16" at 577,349 size 67x20; Text 'Aparente'
   IOField "I/O field_11" at 649,374 size 71x17; FormatPattern 999.99
      ProcessValue <- "VARIAVEIS_QGBT-AUX-01-P100-FP"
      Appearance <- "Digitais_LIT_001-YFS"
   TextField "Text field_17" at 525,371 size 119x20; Text 'Fator de Potência'
   IOField "I/O field_12" at 423,330 size 71x17; FormatPattern 999.99; Unit  A
      ProcessValue <- "VARIAVEIS_QGBT-AUX-01-P100-ITR"
      Appearance <- "Digitais_LIT_001-YFS"
   TextField "Text field_18" at 380,295 size 79x23; Text 'Correntes'
   TextField "Text field_19" at 370,327 size 47x20; Text 'Fase R'
   IOField "I/O field_13" at 423,352 size 71x17; FormatPattern 999.99; Unit  A
      ProcessValue <- "VARIAVEIS_QGBT-AUX-01-P100-ITS"
      Appearance <- "Digitais_LIT_001-YFS"
   TextField "Text field_20" at 371,349 size 46x20; Text 'Fase S'
   IOField "I/O field_15" at 423,374 size 71x17; FormatPattern 999.99; Unit  A
      ProcessValue <- "VARIAVEIS_QGBT-AUX-01-P100-ITT"
      Appearance <- "Digitais_LIT_001-YFS"
   TextField "Text field_21" at 372,371 size 45x20; Text 'Fase T'
   IOField "I/O field_16" at 202,330 size 71x17; FormatPattern 999.99; Unit  V
      ProcessValue <- "VARIAVEIS_QGBT-AUX-01-P100-ETRS"
      Appearance <- "Digitais_LIT_001-YFS"
   TextField "Text field_22" at 166,295 size 66x23; Text 'Tensões'
   TextField "Text field_23" at 133,327 size 63x20; Text 'Fase R/S'
   IOField "I/O field_17" at 202,352 size 71x17; FormatPattern 999.99; Unit  V
      ProcessValue <- "VARIAVEIS_QGBT-AUX-01-P100-ETST"
      Appearance <- "Digitais_LIT_001-YFS"
   TextField "Text field_24" at 133,349 size 61x20; Text 'Fase S/T'
   IOField "I/O field_18" at 202,374 size 71x17; FormatPattern 999.99; Unit  V
      ProcessValue <- "VARIAVEIS_QGBT-AUX-01-P100-ETTR"
      Appearance <- "Digitais_LIT_001-YFS"
   TextField "Text field_25" at 133,371 size 62x20; Text 'Fase T/R'
   TextField "Text field_26" at 350,263 size 120x23; Text 'QGBT-AUX-01'
   IOField "I/O field_6" at 649,154 size 71x17; FormatPattern 999.99; Unit  kW
      ProcessValue <- "VARIAVEIS_PCM-E-CF-01-04-P100-JPT"
      Appearance <- "Digitais_LIT_001-YFS"
   TextField "Text field_9" at 607,119 size 78x23; Text 'Potências'
   TextField "Text field_10" at 604,151 size 40x20; Text 'Ativa'
   IOField "I/O field_7" at 649,176 size 71x17; FormatPattern 999.99; Unit  KVA
      ProcessValue <- "VARIAVEIS_PCM-E-CF-01-04-P100-JST"
      Appearance <- "Digitais_LIT_001-YFS"
   TextField "Text field_11" at 577,173 size 67x20; Text 'Aparente'
   IOField "I/O field_8" at 649,198 size 71x17; FormatPattern 999.99
      ProcessValue <- "VARIAVEIS_PCM-E-CF-01-04-P100-FP"
      Appearance <- "Digitais_LIT_001-YFS"
   TextField "Text field_12" at 525,195 size 119x20; Text 'Fator de Potência'
   IOField "I/O field_3" at 423,154 size 71x17; FormatPattern 999.99; Unit  A
      ProcessValue <- "VARIAVEIS_PCM-E-CF-01-04-P100-ITR"
      Appearance <- "Digitais_LIT_001-YFS"
   TextField "Text field_5" at 380,119 size 79x23; Text 'Correntes'
   TextField "Text field_6" at 370,151 size 47x20; Text 'Fase R'
   IOField "I/O field_4" at 423,176 size 71x17; FormatPattern 999.99; Unit  A
      ProcessValue <- "VARIAVEIS_PCM-E-CF-01-04-P100-ITS"
      Appearance <- "Digitais_LIT_001-YFS"
   TextField "Text field_7" at 371,173 size 46x20; Text 'Fase S'
   IOField "I/O field_5" at 423,198 size 71x17; FormatPattern 999.99; Unit  A
      ProcessValue <- "VARIAVEIS_PCM-E-CF-01-04-P100-ITT"
      Appearance <- "Digitais_LIT_001-YFS"
   TextField "Text field_8" at 372,195 size 45x20; Text 'Fase T'
   IOField "I/O field_14" at 202,154 size 71x17; FormatPattern 999.99; Unit  V
      ProcessValue <- "VARIAVEIS_PCM-E-CF-01-04-P100-ETRS"
      Appearance <- "Digitais_LIT_001-YFS"
   TextField "Text field_1" at 166,119 size 66x23; Text 'Tensões'
   TextField "Text field_2" at 133,151 size 63x20; Text 'Fase R/S'
   IOField "I/O field_1" at 202,176 size 71x17; FormatPattern 999.99; Unit  V
      ProcessValue <- "VARIAVEIS_PCM-E-CF-01-04-P100-ETST"
      Appearance <- "Digitais_LIT_001-YFS"
   TextField "Text field_3" at 133,173 size 61x20; Text 'Fase S/T'
   IOField "I/O field_2" at 202,198 size 71x17; FormatPattern 999.99; Unit  V
      ProcessValue <- "VARIAVEIS_PCM-E-CF-01-04-P100-ETTR"
      Appearance <- "Digitais_LIT_001-YFS"
   TextField "Text field_4" at 133,195 size 62x20; Text 'Fase T/R'
   TextField "Text field_13" at 350,87 size 145x23; Text 'PCM-E-CF-01~04'

screen "Ajustes" 800x480, template "Template_1"
   on GenerateScreen: SetTag("Tag_ScreenNumber", 6)
   TextField "Text field_16" at 164,73 size 135x19; Text 'Setpoints Liga Bombas'
   TextField "Text field_15" at 66,102 size 170x17; Text 'Nivel Liga Bomba Principal (P)'
   TextField "Text field_18" at 66,125 size 225x17; Text 'Nivel Liga Bomba Complementar 1 (C1)'
   IOField "I/O field_3" at 298,98 size 79x21; FormatPattern 99.99; Unit  m
      ProcessValue <- "SETPOINTS_MB-P-SP-L"
   IOField "I/O field_4" at 298,121 size 79x21; FormatPattern 99.99; Unit  m
      ProcessValue <- "SETPOINTS_MB-C1-SP-L"
   TextField "Text field_19" at 66,148 size 225x17; Text 'Nivel Liga Bomba Complementar 2 (C2)'
   TextField "Text field_20" at 66,172 size 225x17; Text 'Nivel Liga Bomba Complementar 3 (C3)'
   IOField "I/O field_5" at 298,144 size 79x21; FormatPattern 99.99; Unit  m
      ProcessValue <- "SETPOINTS_MB-C2-SP-L"
   IOField "I/O field_11" at 298,168 size 79x21; FormatPattern 99.99; Unit  m
      ProcessValue <- "SETPOINTS_MB-C3-SP-L"
   TextField "Text field_21" at 154,379 size 155x17; Text 'Nivel Minimo de Segurança'
   IOField "I/O field_12" at 192,399 size 79x21; FormatPattern 99.99; Unit  m
      ProcessValue <- "SETPOINTS_SP_NVL_MIN"
   TextField "Text field_1" at 66,257 size 175x17; Text 'Nivel Desl. Bomba Principal (P)'
   TextField "Text field_2" at 66,280 size 230x17; Text 'Nivel Desl. Bomba Complementar 1 (C1)'
   IOField "I/O field_1" at 298,253 size 79x21; FormatPattern 99.99; Unit  m
      ProcessValue <- "SETPOINTS_MB-P-SP-DL"
   IOField "I/O field_2" at 298,276 size 79x21; FormatPattern 99.99; Unit  m
      ProcessValue <- "SETPOINTS_MB-C1-SP-DL"
   TextField "Text field_3" at 66,303 size 230x17; Text 'Nivel Desl. Bomba Complementar 2 (C2)'
   TextField "Text field_4" at 66,327 size 230x17; Text 'Nivel Desl. Bomba Complementar 3 (C3)'
   IOField "I/O field_6" at 298,299 size 79x21; FormatPattern 99.99; Unit  m
      ProcessValue <- "SETPOINTS_MB-C2-SP-DL"
   IOField "I/O field_7" at 298,323 size 79x21; FormatPattern 99.99; Unit  m
      ProcessValue <- "SETPOINTS_MB-C3-SP-DL"
   TextField "Text field_5" at 155,225 size 153x19; Text 'Setpoints Desliga Bombas'
   TextField "Text field_6" at 584,144 size 62x19; Text 'Nível EEEB'
   TextField "Text field_7" at 512,179 size 97x17; Text 'Ajuste muito alto'
   TextField "Text field_8" at 548,209 size 61x17; Text 'Ajuste alto'
   IOField "I/O field_8" at 622,177 size 79x21; FormatPattern 999; Unit  %
      ProcessValue <- "SETPOINTS_LIT_001-SPHH"
   IOField "I/O field_9" at 622,207 size 79x21; FormatPattern 999; Unit  %
      ProcessValue <- "SETPOINTS_LIT_001-SPH"
   TextField "Text field_9" at 539,241 size 70x17; Text 'Ajuste baixo'
   TextField "Text field_10" at 503,271 size 106x17; Text 'Ajuste muito baixo'
   IOField "I/O field_10" at 623,239 size 79x21; FormatPattern 999; Unit  %
      ProcessValue <- "SETPOINTS_LIT_001-SPL"
   IOField "I/O field_13" at 623,269 size 79x21; FormatPattern 999; Unit  %
      ProcessValue <- "SETPOINTS_LIT_001-SPLL"
   TextField "Text field_11" at 542,317 size 146x17; Text 'Ajuste nível para controle'
   IOField "I/O field_14" at 576,342 size 79x21; FormatPattern 999; Unit  %
      ProcessValue <- "SETPOINTS_LIT_001-SPC"
   TextField "Text field_12" at 571,73 size 89x19; Text 'Ajustes Gerais'

screen "PID" 800x480, template "Template_1"
   TextField "Text field_6" at 356,57 size 75x19; Text 'PID Bombas'
   IOField "I/O field_10" at 280,105 size 59x17; FormatPattern 9999.999
      ProcessValue <- "PID_PID-EEEB-P"
   IOField "I/O field_8" at 280,129 size 59x17; FormatPattern 9999.999
      ProcessValue <- "PID_PID-EEEB-I"
   IOField "I/O field_13" at 280,153 size 59x17; FormatPattern 9999.999
      ProcessValue <- "PID_PID-EEEB-D"
   IOField "I/O field_15" at 442,105 size 60x17; FormatPattern 999.9; Unit  Hz
      ProcessValue <- "PID_PID-EEEB-MIN"
   IOField "I/O field_16" at 442,129 size 60x17; FormatPattern 999.9; Unit  Hz
      ProcessValue <- "PID_PID-EEEB-MAX"
   IOField "I/O field_17" at 202,81 size 59x17; FormatPattern 999.9; Unit  %
      ProcessValue <- "SETPOINTS_LIT_001-SPC"
   IOField "I/O field_18" at 336,81 size 59x17; FormatPattern 999.9; Unit  %
      ProcessValue <- "VARIAVEIS_LIT_001-P"
   TextField "Text field_21" at 263,81 size 47x16; Text 'Setpoint'
   TextField "Text field_1" at 398,81 size 47x16; Text 'Medição'
   IOField "I/O field_1" at 442,153 size 59x17; FormatPattern 999.9; Unit  %
      ProcessValue <- "PID_PID-EEEB-DB"
   IOField "I/O field_2" at 471,81 size 59x17; FormatPattern 999.9; Unit  %
      ProcessValue <- "PID_PID-EEEB-VR"
   TextField "Text field_2" at 534,81 size 79x16; Text 'Valor Relativo'
   TextField "Text field_3" at 341,106 size 71x16; Text 'Proporcional'
   TextField "Text field_4" at 341,130 size 44x16; Text 'Integral'
   TextField "Text field_5" at 341,154 size 56x16; Text 'Derivativa'
   TextField "Text field_7" at 504,106 size 97x16; Text 'CV Minimo Saida'
   TextField "Text field_8" at 504,130 size 100x16; Text 'CV Maximo Saida'
   TextField "Text field_9" at 504,154 size 72x16; Text 'Banda Morta'
   TrendView "Trend view_1" at 0,174 size 799x267
   Button "Button_5" at 254,106 size 19x17; TextOff 'P'; Authorization "Operate"
      on Press: InvertBit("COMANDOS_PID-EEEB-HP")
      Appearance <- "COMANDOS_PID-EEEB-HP"
   Button "Button_1" at 254,129 size 19x17; TextOff 'I'; Authorization "Operate"
      on Press: InvertBit("COMANDOS_PID-EEEB-HI")
      Appearance <- "COMANDOS_PID-EEEB-HI"
   Button "Button_2" at 254,153 size 19x17; TextOff 'D'; Authorization "Operate"
      on Press: InvertBit("COMANDOS_PID-EEEB-HD")
      Appearance <- "COMANDOS_PID-EEEB-HD"
   TextField "Text field_10" at 149,106 size 101x16; Text 'Hab. Proporcional'
   TextField "Text field_11" at 149,130 size 74x16; Text 'Hab. Integral'
   TextField "Text field_12" at 149,154 size 86x16; Text 'Hab. Derivativa'

screen "Comandos" 800x480, template "Template_1"
   TextField "Text field_6" at 237,71 size 99x19; Text 'Comando MB-01'
   Button "Button_5" at 209,136 size 70x30; TextOff 'Automático'; Authorization "Operate"
      on Press: SetBit("COMANDOS_MB-01-HS1")
      Appearance <- "COMANDOS_MB-01-HS1"
   Button "Button_8" at 295,136 size 70x30; TextOff 'Manual'; Authorization "Operate"
      on Press: ResetBit("COMANDOS_MB-01-HS1")
      Appearance <- "COMANDOS_MB-01-HS1"
   Button "Button_1" at 209,174 size 70x30; TextOff 'Liga'; Authorization "Operate"
      on Press: SetBit("COMANDOS_MB-01-HS2")
   Button "Button_2" at 295,174 size 70x30; TextOff 'Desliga'; Authorization "Operate"
      on Press: SetBit("COMANDOS_MB-01-HS3")
   TextField "Text field_7" at 199,104 size 118x17; Text 'Ajuste de velocidade'
   IOField "I/O field_10" at 322,100 size 79x21; FormatPattern 99.99; Unit  Hz
      ProcessValue <- "SETPOINTS_MB-01-SP"
   Button "Button_3" at 295,212 size 70x30; TextOff 'Reset'; Authorization "Operate"
      on Press: SetBit("COMANDOS_MB-01-HS4")
   TextField "Text field_8" at 482,71 size 99x19; Text 'Comando MB-02'
   Button "Button_4" at 454,136 size 70x30; TextOff 'Automático'; Authorization "Operate"
      on Press: SetBit("COMANDOS_MB-02-HS1")
      Appearance <- "COMANDOS_MB-02-HS1"
   Button "Button_6" at 540,136 size 70x30; TextOff 'Manual'; Authorization "Operate"
      on Press: ResetBit("COMANDOS_MB-02-HS1")
      Appearance <- "COMANDOS_MB-02-HS1"
   Button "Button_7" at 454,174 size 70x30; TextOff 'Liga'; Authorization "Operate"
      on Press: SetBit("COMANDOS_MB-02-HS2")
   Button "Button_9" at 540,174 size 70x30; TextOff 'Desliga'; Authorization "Operate"
      on Press: SetBit("COMANDOS_MB-02-HS3")
   TextField "Text field_9" at 442,104 size 118x17; Text 'Ajuste de velocidade'
   IOField "I/O field_8" at 564,100 size 79x21; FormatPattern 99.99; Unit  Hz
      ProcessValue <- "SETPOINTS_MB-02-SP"
   Button "Button_10" at 540,212 size 70x30; TextOff 'Reset'; Authorization "Operate"
      on Press: SetBit("COMANDOS_MB-02-HS4")
   TextField "Text field_10" at 237,259 size 99x19; Text 'Comando MB-03'
   Button "Button_11" at 209,324 size 70x30; TextOff 'Automático'; Authorization "Operate"
      on Press: SetBit("COMANDOS_MB-03-HS1")
      Appearance <- "COMANDOS_MB-03-HS1"
   Button "Button_12" at 295,324 size 70x30; TextOff 'Manual'; Authorization "Operate"
      on Press: ResetBit("COMANDOS_MB-03-HS1")
      Appearance <- "COMANDOS_MB-03-HS1"
   Button "Button_13" at 209,362 size 70x30; TextOff 'Liga'; Authorization "Operate"
      on Press: SetBit("COMANDOS_MB-03-HS2")
   Button "Button_14" at 295,362 size 70x30; TextOff 'Desliga'; Authorization "Operate"
      on Press: SetBit("COMANDOS_MB-03-HS3")
   TextField "Text field_11" at 199,292 size 118x17; Text 'Ajuste de velocidade'
   IOField "I/O field_9" at 322,288 size 79x21; FormatPattern 99.99; Unit  Hz
      ProcessValue <- "SETPOINTS_MB-03-SP"
   Button "Button_15" at 295,400 size 70x30; TextOff 'Reset'; Authorization "Operate"
      on Press: SetBit("COMANDOS_MB-03-HS4")
   TextField "Text field_12" at 482,259 size 99x19; Text 'Comando MB-04'
   Button "Button_16" at 454,324 size 70x30; TextOff 'Automático'; Authorization "Operate"
      on Press: SetBit("COMANDOS_MB-04-HS1")
      Appearance <- "COMANDOS_MB-04-HS1"
   Button "Button_17" at 540,324 size 70x30; TextOff 'Manual'; Authorization "Operate"
      on Press: ResetBit("COMANDOS_MB-04-HS1")
      Appearance <- "COMANDOS_MB-04-HS1"
   Button "Button_18" at 454,362 size 70x30; TextOff 'Liga'; Authorization "Operate"
      on Press: SetBit("COMANDOS_MB-04-HS2")
   Button "Button_19" at 540,362 size 70x30; TextOff 'Desliga'; Authorization "Operate"
      on Press: SetBit("COMANDOS_MB-04-HS3")
   TextField "Text field_13" at 442,292 size 118x17; Text 'Ajuste de velocidade'
   IOField "I/O field_13" at 564,288 size 79x21; FormatPattern 99.99; Unit  Hz
      ProcessValue <- "SETPOINTS_MB-04-SP"
   Button "Button_20" at 540,400 size 70x30; TextOff 'Reset'; Authorization "Operate"
      on Press: SetBit("COMANDOS_MB-04-HS4")
*)